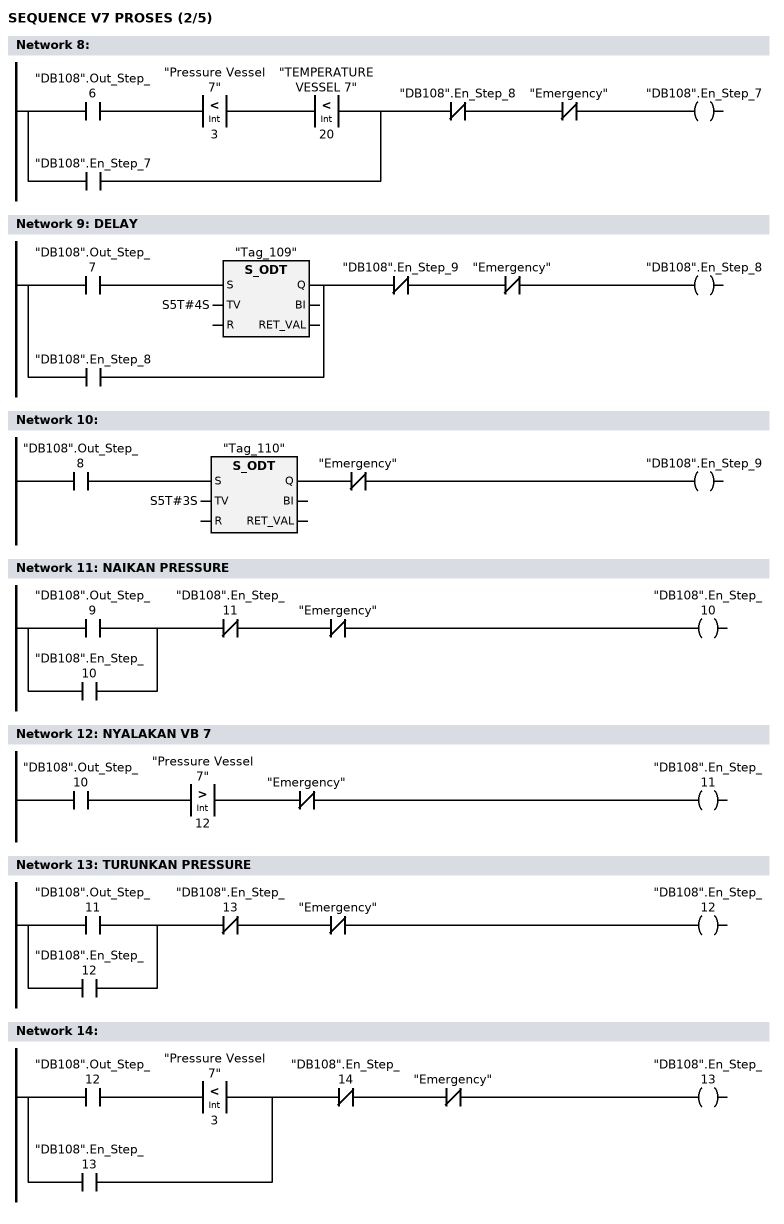
   RUNG wire#powerrail
      Contact( "DB108".Out_Step_6 )
      { S7_Templates := "SrcType := Int" } LT_Contact(in1 := "Pressure Vessel 7", in2 := 3)
      { S7_Templates := "SrcType := Int" } LT_Contact(in1 := "TEMPERATURE VESSEL 7", in2 := 20)
      wire#w1
      I_Contact( "DB108".En_Step_8 )
      I_Contact( "Emergency" )
      Coil( "DB108".En_Step_7 )
   END_RUNG
   RUNG wire#powerrail
      Contact( "DB108".En_Step_7 )
   END_RUNG wire#w1
   // the same network as SCL:
   "DB108".En_Step_7 := (("DB108".Out_Step_6 AND ("Pressure Vessel 7" < 3) AND ("TEMPERATURE VESSEL 7" < 20)) OR "DB108".En_Step_7) AND NOT "DB108".En_Step_8 AND NOT "Emergency";
END_REGION

REGION Network 9: DELAY
   RUNG wire#powerrail
      Contact( "DB108".Out_Step_7 )
      S_ODT(T_NO := "Tag_109", TV := S5T#4S, R :=, BI =>, RET_VAL =>)
      wire#w1
      I_Contact( "DB108".En_Step_9 )
      I_Contact( "Emergency" )
      Coil( "DB108".En_Step_8 )
   END_RUNG
   RUNG wire#powerrail
      Contact( "DB108".En_Step_8 )
   END_RUNG wire#w1
   // the same network as SCL:
   #_s5time1 := S_ODT(T_NO := "Tag_109", S := "DB108".Out_Step_7, TV := S5T#4S, Q => #_w1);
   "DB108".En_Step_8 := (#_w1 OR "DB108".En_Step_8) AND NOT "DB108".En_Step_9 AND NOT "Emergency";
END_REGION

REGION Network 10
   RUNG wire#powerrail
      Contact( "DB108".Out_Step_8 )
      S_ODT(T_NO := "Tag_110", TV := S5T#3S, R :=, BI =>, RET_VAL =>)
      I_Contact( "Emergency" )
      Coil( "DB108".En_Step_9 )
   END_RUNG
   // the same network as SCL:
   #_s5time1 := S_ODT(T_NO := "Tag_110", S := "DB108".Out_Step_8, TV := S5T#3S, Q => #_w1);
   "DB108".En_Step_9 := #_w1 AND NOT "Emergency";
END_REGION

REGION Network 11: NAIKAN PRESSURE
   RUNG wire#powerrail
      Contact( "DB108".Out_Step_9 )
      wire#w1
      I_Contact( "DB108".En_Step_11 )
      I_Contact( "Emergency" )
      Coil( "DB108".En_Step_10 )
   END_RUNG
   RUNG wire#powerrail
      Contact( "DB108".En_Step_10 )
   END_RUNG wire#w1
   // the same network as SCL:
   "DB108".En_Step_10 := ("DB108".Out_Step_9 OR "DB108".En_Step_10) AND NOT "DB108".En_Step_11 AND NOT "Emergency";
END_REGION

REGION Network 12: NYALAKAN VB 7
   RUNG wire#powerrail
      Contact( "DB108".Out_Step_10 )
      { S7_Templates := "SrcType := Int" } GT_Contact(in1 := "Pressure Vessel 7", in2 := 12)
      I_Contact( "Emergency" )
      Coil( "DB108".En_Step_11 )
   END_RUNG
   // the same network as SCL:
   "DB108".En_Step_11 := "DB108".Out_Step_10 AND ("Pressure Vessel 7" > 12) AND NOT "Emergency";
END_REGION

REGION Network 13: TURUNKAN PRESSURE
   RUNG wire#powerrail
      Contact( "DB108".Out_Step_11 )
      wire#w1
      I_Contact( "DB108".En_Step_13 )
      I_Contact( "Emergency" )
      Coil( "DB108".En_Step_12 )
   END_RUNG
   RUNG wire#powerrail
      Contact( "DB108".En_Step_12 )
   END_RUNG wire#w1
   // the same network as SCL:
   "DB108".En_Step_12 := ("DB108".Out_Step_11 OR "DB108".En_Step_12) AND NOT "DB108".En_Step_13 AND NOT "Emergency";
END_REGION

REGION Network 14
   RUNG wire#powerrail
      Contact( "DB108".Out_Step_12 )
      { S7_Templates := "SrcType := Int" } LT_Contact(in1 := "Pressure Vessel 7", in2 := 3)
      wire#w1
      I_Contact( "DB108".En_Step_14 )
      I_Contact( "Emergency" )
      Coil( "DB108".En_Step_13 )
   END_RUNG
   RUNG wire#powerrail
      Contact( "DB108".En_Step_13 )
   END_RUNG wire#w1
   // the same network as SCL:
   "DB108".En_Step_13 := (("DB108".Out_Step_12 AND ("Pressure Vessel 7" < 3)) OR "DB108".En_Step_13) AND NOT "DB108".En_Step_14 AND NOT "Emergency";
END_REGION

REGION Network 15
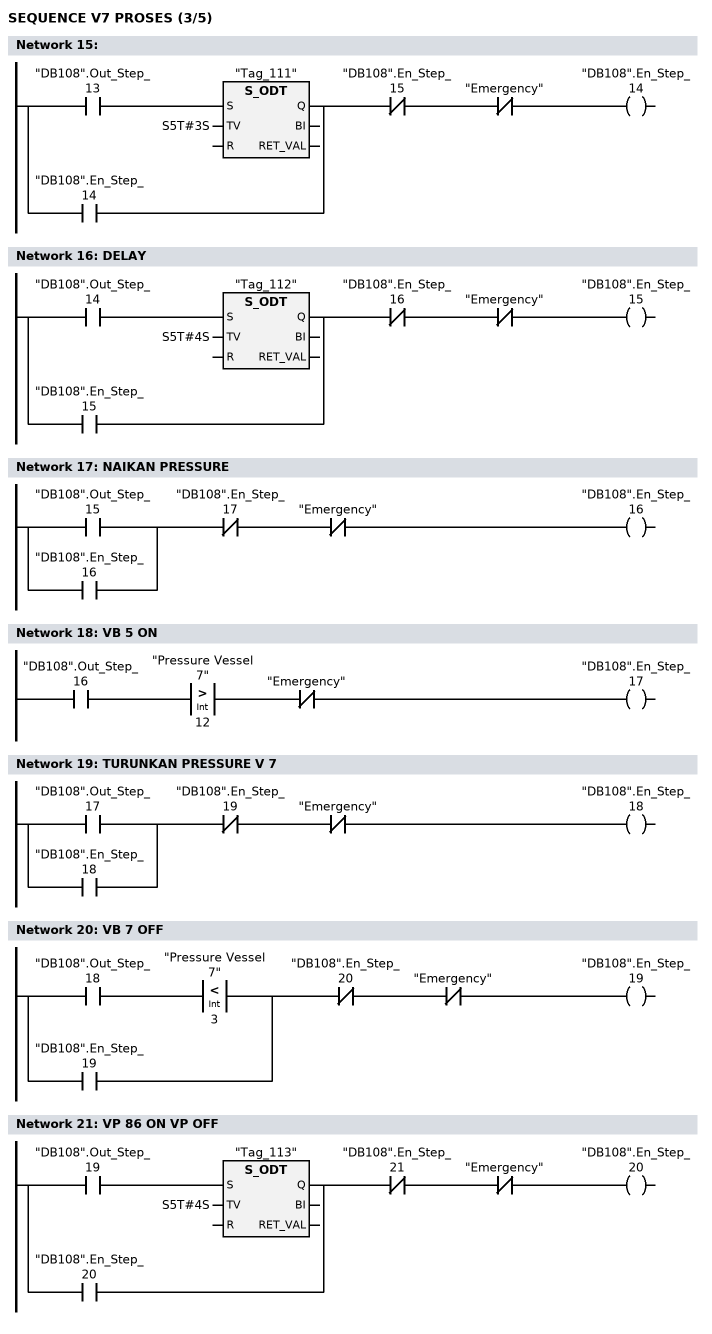
   RUNG wire#powerrail
      Contact( "DB108".Out_Step_13 )
      S_ODT(T_NO := "Tag_111", TV := S5T#3S, R :=, BI =>, RET_VAL =>)
      wire#w1
      I_Contact( "DB108".En_Step_15 )
      I_Contact( "Emergency" )
      Coil( "DB108".En_Step_14 )
   END_RUNG
   RUNG wire#powerrail
      Contact( "DB108".En_Step_14 )
   END_RUNG wire#w1
   // the same network as SCL:
   #_s5time1 := S_ODT(T_NO := "Tag_111", S := "DB108".Out_Step_13, TV := S5T#3S, Q => #_w1);
   "DB108".En_Step_14 := (#_w1 OR "DB108".En_Step_14) AND NOT "DB108".En_Step_15 AND NOT "Emergency";
END_REGION

REGION Network 16: DELAY
   RUNG wire#powerrail
      Contact( "DB108".Out_Step_14 )
      S_ODT(T_NO := "Tag_112", TV := S5T#4S, R :=, BI =>, RET_VAL =>)
      wire#w1
      I_Contact( "DB108".En_Step_16 )
      I_Contact( "Emergency" )
      Coil( "DB108".En_Step_15 )
   END_RUNG
   RUNG wire#powerrail
      Contact( "DB108".En_Step_15 )
   END_RUNG wire#w1
   // the same network as SCL:
   #_s5time1 := S_ODT(T_NO := "Tag_112", S := "DB108".Out_Step_14, TV := S5T#4S, Q => #_w1);
   "DB108".En_Step_15 := (#_w1 OR "DB108".En_Step_15) AND NOT "DB108".En_Step_16 AND NOT "Emergency";
END_REGION

REGION Network 17: NAIKAN PRESSURE
   RUNG wire#powerrail
      Contact( "DB108".Out_Step_15 )
      wire#w1
      I_Contact( "DB108".En_Step_17 )
      I_Contact( "Emergency" )
      Coil( "DB108".En_Step_16 )
   END_RUNG
   RUNG wire#powerrail
      Contact( "DB108".En_Step_16 )
   END_RUNG wire#w1
   // the same network as SCL:
   "DB108".En_Step_16 := ("DB108".Out_Step_15 OR "DB108".En_Step_16) AND NOT "DB108".En_Step_17 AND NOT "Emergency";
END_REGION

REGION Network 18: VB 5 ON
   RUNG wire#powerrail
      Contact( "DB108".Out_Step_16 )
      { S7_Templates := "SrcType := Int" } GT_Contact(in1 := "Pressure Vessel 7", in2 := 12)
      I_Contact( "Emergency" )
      Coil( "DB108".En_Step_17 )
   END_RUNG
   // the same network as SCL:
   "DB108".En_Step_17 := "DB108".Out_Step_16 AND ("Pressure Vessel 7" > 12) AND NOT "Emergency";
END_REGION

REGION Network 19: TURUNKAN PRESSURE V 7
   RUNG wire#powerrail
      Contact( "DB108".Out_Step_17 )
      wire#w1
      I_Contact( "DB108".En_Step_19 )
      I_Contact( "Emergency" )
      Coil( "DB108".En_Step_18 )
   END_RUNG
   RUNG wire#powerrail
      Contact( "DB108".En_Step_18 )
   END_RUNG wire#w1
   // the same network as SCL:
   "DB108".En_Step_18 := ("DB108".Out_Step_17 OR "DB108".En_Step_18) AND NOT "DB108".En_Step_19 AND NOT "Emergency";
END_REGION

REGION Network 20: VB 7 OFF
   RUNG wire#powerrail
      Contact( "DB108".Out_Step_18 )
      { S7_Templates := "SrcType := Int" } LT_Contact(in1 := "Pressure Vessel 7", in2 := 3)
      wire#w1
      I_Contact( "DB108".En_Step_20 )
      I_Contact( "Emergency" )
      Coil( "DB108".En_Step_19 )
   END_RUNG
   RUNG wire#powerrail
      Contact( "DB108".En_Step_19 )
   END_RUNG wire#w1
   // the same network as SCL:
   "DB108".En_Step_19 := (("DB108".Out_Step_18 AND ("Pressure Vessel 7" < 3)) OR "DB108".En_Step_19) AND NOT "DB108".En_Step_20 AND NOT "Emergency";
END_REGION

REGION Network 21: VP 86 ON VP OFF
   RUNG wire#powerrail
      Contact( "DB108".Out_Step_19 )
      S_ODT(T_NO := "Tag_113", TV := S5T#4S, R :=, BI =>, RET_VAL =>)
      wire#w1
      I_Contact( "DB108".En_Step_21 )
      I_Contact( "Emergency" )
      Coil( "DB108".En_Step_20 )
   END_RUNG
   RUNG wire#powerrail
      Contact( "DB108".En_Step_20 )
   END_RUNG wire#w1
   // the same network as SCL:
   #_s5time1 := S_ODT(T_NO := "Tag_113", S := "DB108".Out_Step_19, TV := S5T#4S, Q => #_w1);
   "DB108".En_Step_20 := (#_w1 OR "DB108".En_Step_20) AND NOT "DB108".En_Step_21 AND NOT "Emergency";
END_REGION

REGION Network 22: VP 86 OFF VP 87 ON
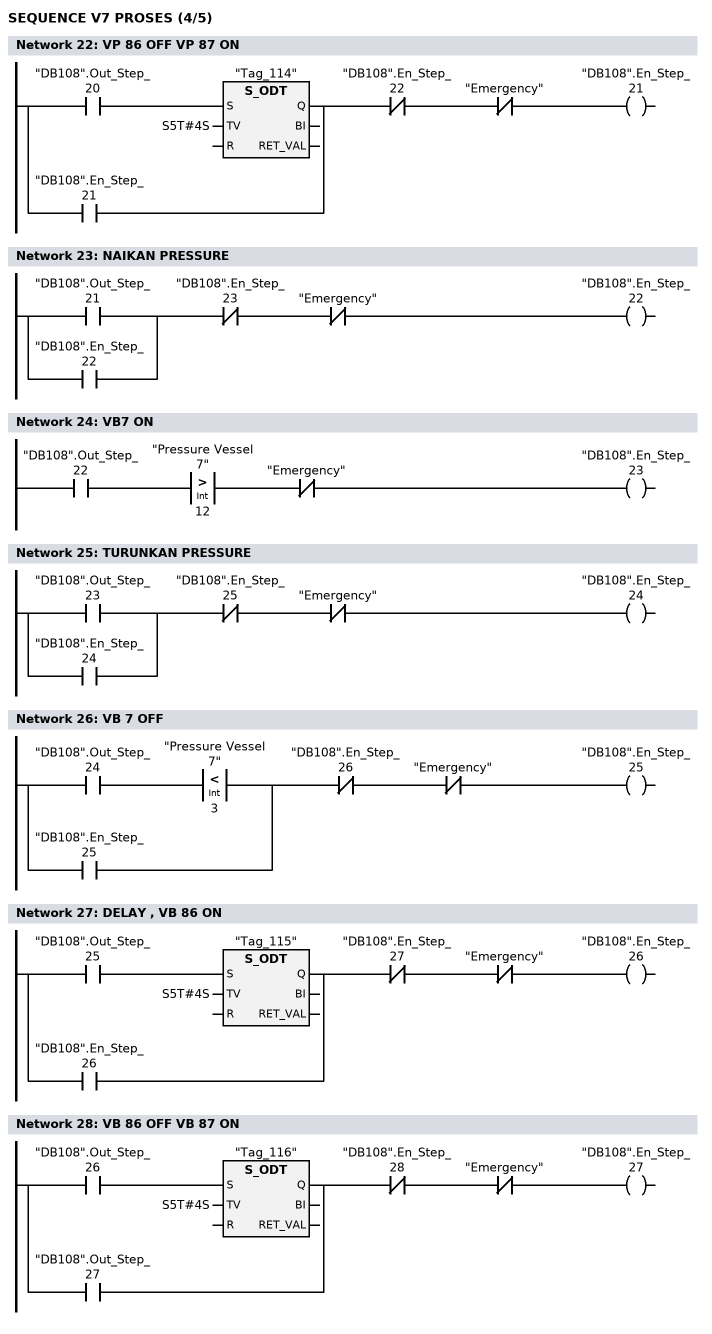
   RUNG wire#powerrail
      Contact( "DB108".Out_Step_20 )
      S_ODT(T_NO := "Tag_114", TV := S5T#4S, R :=, BI =>, RET_VAL =>)
      wire#w1
      I_Contact( "DB108".En_Step_22 )
      I_Contact( "Emergency" )
      Coil( "DB108".En_Step_21 )
   END_RUNG
   RUNG wire#powerrail
      Contact( "DB108".En_Step_21 )
   END_RUNG wire#w1
   // the same network as SCL:
   #_s5time1 := S_ODT(T_NO := "Tag_114", S := "DB108".Out_Step_20, TV := S5T#4S, Q => #_w1);
   "DB108".En_Step_21 := (#_w1 OR "DB108".En_Step_21) AND NOT "DB108".En_Step_22 AND NOT "Emergency";
END_REGION

REGION Network 23: NAIKAN PRESSURE
   RUNG wire#powerrail
      Contact( "DB108".Out_Step_21 )
      wire#w1
      I_Contact( "DB108".En_Step_23 )
      I_Contact( "Emergency" )
      Coil( "DB108".En_Step_22 )
   END_RUNG
   RUNG wire#powerrail
      Contact( "DB108".En_Step_22 )
   END_RUNG wire#w1
   // the same network as SCL:
   "DB108".En_Step_22 := ("DB108".Out_Step_21 OR "DB108".En_Step_22) AND NOT "DB108".En_Step_23 AND NOT "Emergency";
END_REGION

REGION Network 24: VB7 ON
   RUNG wire#powerrail
      Contact( "DB108".Out_Step_22 )
      { S7_Templates := "SrcType := Int" } GT_Contact(in1 := "Pressure Vessel 7", in2 := 12)
      I_Contact( "Emergency" )
      Coil( "DB108".En_Step_23 )
   END_RUNG
   // the same network as SCL:
   "DB108".En_Step_23 := "DB108".Out_Step_22 AND ("Pressure Vessel 7" > 12) AND NOT "Emergency";
END_REGION

REGION Network 25: TURUNKAN PRESSURE
   RUNG wire#powerrail
      Contact( "DB108".Out_Step_23 )
      wire#w1
      I_Contact( "DB108".En_Step_25 )
      I_Contact( "Emergency" )
      Coil( "DB108".En_Step_24 )
   END_RUNG
   RUNG wire#powerrail
      Contact( "DB108".En_Step_24 )
   END_RUNG wire#w1
   // the same network as SCL:
   "DB108".En_Step_24 := ("DB108".Out_Step_23 OR "DB108".En_Step_24) AND NOT "DB108".En_Step_25 AND NOT "Emergency";
END_REGION

REGION Network 26: VB 7 OFF
   RUNG wire#powerrail
      Contact( "DB108".Out_Step_24 )
      { S7_Templates := "SrcType := Int" } LT_Contact(in1 := "Pressure Vessel 7", in2 := 3)
      wire#w1
      I_Contact( "DB108".En_Step_26 )
      I_Contact( "Emergency" )
      Coil( "DB108".En_Step_25 )
   END_RUNG
   RUNG wire#powerrail
      Contact( "DB108".En_Step_25 )
   END_RUNG wire#w1
   // the same network as SCL:
   "DB108".En_Step_25 := (("DB108".Out_Step_24 AND ("Pressure Vessel 7" < 3)) OR "DB108".En_Step_25) AND NOT "DB108".En_Step_26 AND NOT "Emergency";
END_REGION

REGION Network 27: DELAY , VB 86 ON
   RUNG wire#powerrail
      Contact( "DB108".Out_Step_25 )
      S_ODT(T_NO := "Tag_115", TV := S5T#4S, R :=, BI =>, RET_VAL =>)
      wire#w1
      I_Contact( "DB108".En_Step_27 )
      I_Contact( "Emergency" )
      Coil( "DB108".En_Step_26 )
   END_RUNG
   RUNG wire#powerrail
      Contact( "DB108".En_Step_26 )
   END_RUNG wire#w1
   // the same network as SCL:
   #_s5time1 := S_ODT(T_NO := "Tag_115", S := "DB108".Out_Step_25, TV := S5T#4S, Q => #_w1);
   "DB108".En_Step_26 := (#_w1 OR "DB108".En_Step_26) AND NOT "DB108".En_Step_27 AND NOT "Emergency";
END_REGION

REGION Network 28: VB 86 OFF VB 87 ON
   RUNG wire#powerrail
      Contact( "DB108".Out_Step_26 )
      S_ODT(T_NO := "Tag_116", TV := S5T#4S, R :=, BI =>, RET_VAL =>)
      wire#w1
      I_Contact( "DB108".En_Step_28 )
      I_Contact( "Emergency" )
      Coil( "DB108".En_Step_27 )
   END_RUNG
   RUNG wire#powerrail
      Contact( "DB108".Out_Step_27 )
   END_RUNG wire#w1
   // the same network as SCL:
   #_s5time1 := S_ODT(T_NO := "Tag_116", S := "DB108".Out_Step_26, TV := S5T#4S, Q => #_w1);
   "DB108".En_Step_27 := (#_w1 OR "DB108".Out_Step_27) AND NOT "DB108".En_Step_28 AND NOT "Emergency";
END_REGION

REGION Network 29
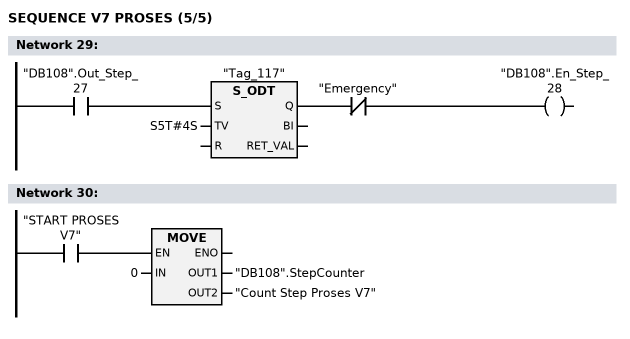
   RUNG wire#powerrail
      Contact( "DB108".Out_Step_27 )
      S_ODT(T_NO := "Tag_117", TV := S5T#4S, R :=, BI =>, RET_VAL =>)
      I_Contact( "Emergency" )
      Coil( "DB108".En_Step_28 )
   END_RUNG
   // the same network as SCL:
   #_s5time1 := S_ODT(T_NO := "Tag_117", S := "DB108".Out_Step_27, TV := S5T#4S, Q => #_w1);
   "DB108".En_Step_28 := #_w1 AND NOT "Emergency";
END_REGION

REGION Network 30
   RUNG wire#powerrail
      Contact( "START PROSES V7" )
      Move(in := 0, out1 => "DB108".StepCounter, out2 => "Count Step Proses V7")
   END_RUNG
   // the same network as SCL:
   IF "START PROSES V7" THEN
       "DB108".StepCounter := 0;
       "Count Step Proses V7" := 0;
   END_IF;
END_REGION
END_FUNCTION

FUNCTION "SEQUENCE V2 PREPARATION" : Void   // FC23, LAD
{ S7_Optimized_Access := 'TRUE' }
VERSION : 0.1
   VAR_TEMP   // added for the SCL form of the ladder/FBD networks
      _w1 : Bool;
      _s5time1 : S5Time;
      _w2 : Bool;
      _s5time2 : S5Time;
   END_VAR
BEGIN

REGION Network 1: Start Preparation
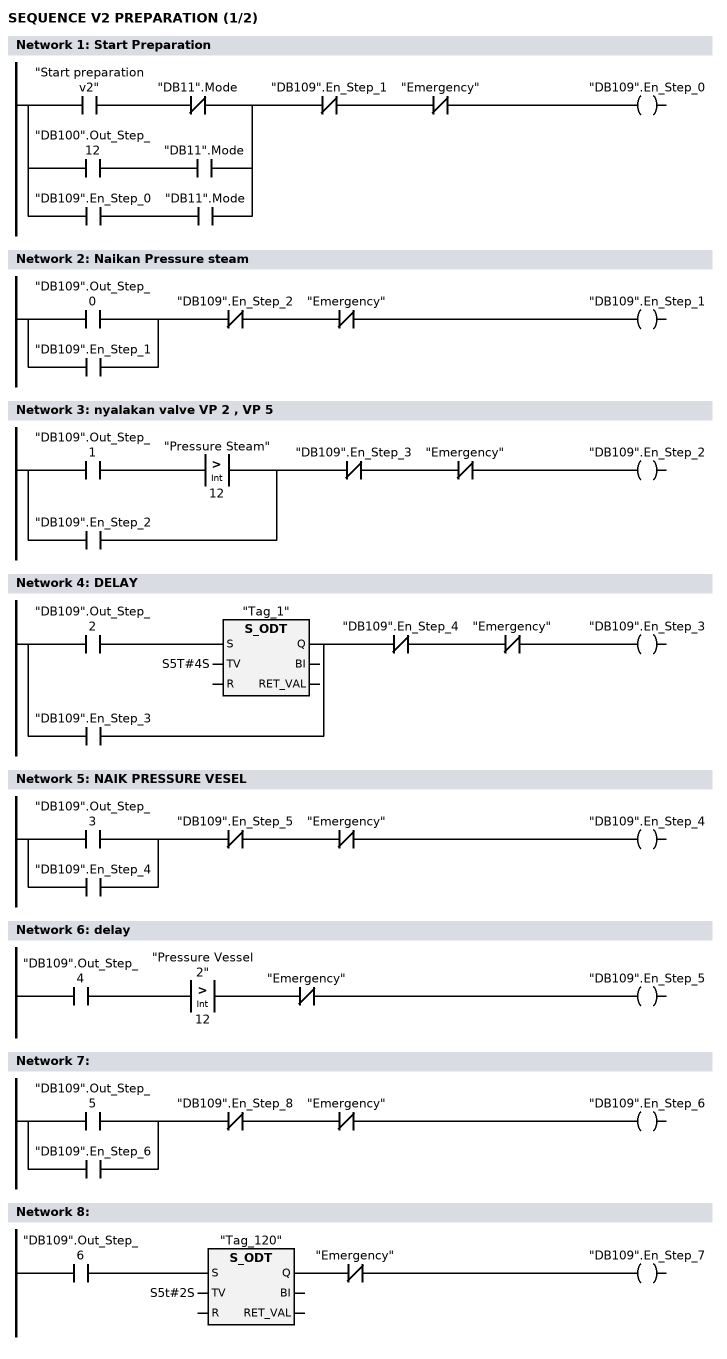
   RUNG wire#powerrail
      Contact( "Start preparation v2" )
      I_Contact( "DB11".Mode )
      wire#w1
      I_Contact( "DB109".En_Step_1 )
      I_Contact( "Emergency" )
      Coil( "DB109".En_Step_0 )
   END_RUNG
   RUNG wire#powerrail
      Contact( "DB100".Out_Step_12 )
      Contact( "DB11".Mode )
   END_RUNG wire#w1
   RUNG wire#powerrail
      Contact( "DB109".En_Step_0 )
      Contact( "DB11".Mode )
   END_RUNG wire#w1
   // the same network as SCL:
   "DB109".En_Step_0 := (("Start preparation v2" AND NOT "DB11".Mode) OR ("DB100".Out_Step_12 AND "DB11".Mode) OR ("DB109".En_Step_0 AND "DB11".Mode)) AND NOT "DB109".En_Step_1 AND NOT "Emergency";
END_REGION

REGION Network 2: Naikan Pressure steam
   RUNG wire#powerrail
      Contact( "DB109".Out_Step_0 )
      wire#w1
      I_Contact( "DB109".En_Step_2 )
      I_Contact( "Emergency" )
      Coil( "DB109".En_Step_1 )
   END_RUNG
   RUNG wire#powerrail
      Contact( "DB109".En_Step_1 )
   END_RUNG wire#w1
   // the same network as SCL:
   "DB109".En_Step_1 := ("DB109".Out_Step_0 OR "DB109".En_Step_1) AND NOT "DB109".En_Step_2 AND NOT "Emergency";
END_REGION

REGION Network 3: nyalakan valve VP 2 , VP 5
   RUNG wire#powerrail
      Contact( "DB109".Out_Step_1 )
      { S7_Templates := "SrcType := Int" } GT_Contact(in1 := "Pressure Steam", in2 := 12)
      wire#w1
      I_Contact( "DB109".En_Step_3 )
      I_Contact( "Emergency" )
      Coil( "DB109".En_Step_2 )
   END_RUNG
   RUNG wire#powerrail
      Contact( "DB109".En_Step_2 )
   END_RUNG wire#w1
   // the same network as SCL:
   "DB109".En_Step_2 := (("DB109".Out_Step_1 AND ("Pressure Steam" > 12)) OR "DB109".En_Step_2) AND NOT "DB109".En_Step_3 AND NOT "Emergency";
END_REGION

REGION Network 4: DELAY
   RUNG wire#powerrail
      Contact( "DB109".Out_Step_2 )
      S_ODT(T_NO := "Tag_1", TV := S5T#4S, R :=, BI =>, RET_VAL =>)
      wire#w1
      I_Contact( "DB109".En_Step_4 )
      I_Contact( "Emergency" )
      Coil( "DB109".En_Step_3 )
   END_RUNG
   RUNG wire#powerrail
      Contact( "DB109".En_Step_3 )
   END_RUNG wire#w1
   // the same network as SCL:
   #_s5time1 := S_ODT(T_NO := "Tag_1", S := "DB109".Out_Step_2, TV := S5T#4S, Q => #_w1);
   "DB109".En_Step_3 := (#_w1 OR "DB109".En_Step_3) AND NOT "DB109".En_Step_4 AND NOT "Emergency";
END_REGION

REGION Network 5: NAIK PRESSURE VESEL
   RUNG wire#powerrail
      Contact( "DB109".Out_Step_3 )
      wire#w1
      I_Contact( "DB109".En_Step_5 )
      I_Contact( "Emergency" )
      Coil( "DB109".En_Step_4 )
   END_RUNG
   RUNG wire#powerrail
      Contact( "DB109".En_Step_4 )
   END_RUNG wire#w1
   // the same network as SCL:
   "DB109".En_Step_4 := ("DB109".Out_Step_3 OR "DB109".En_Step_4) AND NOT "DB109".En_Step_5 AND NOT "Emergency";
END_REGION

REGION Network 6: delay
   RUNG wire#powerrail
      Contact( "DB109".Out_Step_4 )
      { S7_Templates := "SrcType := Int" } GT_Contact(in1 := "Pressure Vessel 2", in2 := 12)
      I_Contact( "Emergency" )
      Coil( "DB109".En_Step_5 )
   END_RUNG
   // the same network as SCL:
   "DB109".En_Step_5 := "DB109".Out_Step_4 AND ("Pressure Vessel 2" > 12) AND NOT "Emergency";
END_REGION

REGION Network 7
   RUNG wire#powerrail
      Contact( "DB109".Out_Step_5 )
      wire#w1
      I_Contact( "DB109".En_Step_8 )
      I_Contact( "Emergency" )
      Coil( "DB109".En_Step_6 )
   END_RUNG
   RUNG wire#powerrail
      Contact( "DB109".En_Step_6 )
   END_RUNG wire#w1
   // the same network as SCL:
   "DB109".En_Step_6 := ("DB109".Out_Step_5 OR "DB109".En_Step_6) AND NOT "DB109".En_Step_8 AND NOT "Emergency";
END_REGION

REGION Network 8
   RUNG wire#powerrail
      Contact( "DB109".Out_Step_6 )
      S_ODT(T_NO := "Tag_120", TV := S5t#2S, R :=, BI =>, RET_VAL =>)
      I_Contact( "Emergency" )
      Coil( "DB109".En_Step_7 )
   END_RUNG
   // the same network as SCL:
   #_s5time1 := S_ODT(T_NO := "Tag_120", S := "DB109".Out_Step_6, TV := S5t#2S, Q => #_w1);
   "DB109".En_Step_7 := #_w1 AND NOT "Emergency";
END_REGION

REGION Network 9: TURUNKAN PRESSURE
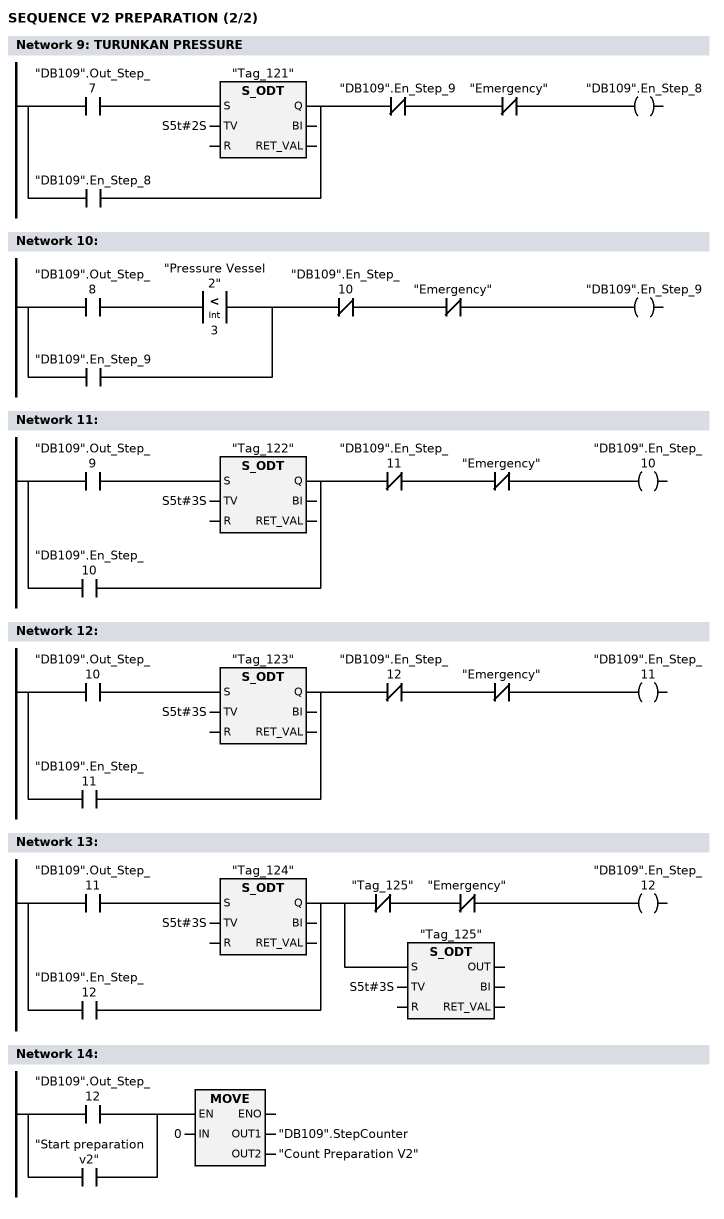
   RUNG wire#powerrail
      Contact( "DB109".Out_Step_7 )
      S_ODT(T_NO := "Tag_121", TV := S5t#2S, R :=, BI =>, RET_VAL =>)
      wire#w1
      I_Contact( "DB109".En_Step_9 )
      I_Contact( "Emergency" )
      Coil( "DB109".En_Step_8 )
   END_RUNG
   RUNG wire#powerrail
      Contact( "DB109".En_Step_8 )
   END_RUNG wire#w1
   // the same network as SCL:
   #_s5time1 := S_ODT(T_NO := "Tag_121", S := "DB109".Out_Step_7, TV := S5t#2S, Q => #_w1);
   "DB109".En_Step_8 := (#_w1 OR "DB109".En_Step_8) AND NOT "DB109".En_Step_9 AND NOT "Emergency";
END_REGION

REGION Network 10
   RUNG wire#powerrail
      Contact( "DB109".Out_Step_8 )
      { S7_Templates := "SrcType := Int" } LT_Contact(in1 := "Pressure Vessel 2", in2 := 3)
      wire#w1
      I_Contact( "DB109".En_Step_10 )
      I_Contact( "Emergency" )
      Coil( "DB109".En_Step_9 )
   END_RUNG
   RUNG wire#powerrail
      Contact( "DB109".En_Step_9 )
   END_RUNG wire#w1
   // the same network as SCL:
   "DB109".En_Step_9 := (("DB109".Out_Step_8 AND ("Pressure Vessel 2" < 3)) OR "DB109".En_Step_9) AND NOT "DB109".En_Step_10 AND NOT "Emergency";
END_REGION

REGION Network 11
   RUNG wire#powerrail
      Contact( "DB109".Out_Step_9 )
      S_ODT(T_NO := "Tag_122", TV := S5t#3S, R :=, BI =>, RET_VAL =>)
      wire#w1
      I_Contact( "DB109".En_Step_11 )
      I_Contact( "Emergency" )
      Coil( "DB109".En_Step_10 )
   END_RUNG
   RUNG wire#powerrail
      Contact( "DB109".En_Step_10 )
   END_RUNG wire#w1
   // the same network as SCL:
   #_s5time1 := S_ODT(T_NO := "Tag_122", S := "DB109".Out_Step_9, TV := S5t#3S, Q => #_w1);
   "DB109".En_Step_10 := (#_w1 OR "DB109".En_Step_10) AND NOT "DB109".En_Step_11 AND NOT "Emergency";
END_REGION

REGION Network 12
   RUNG wire#powerrail
      Contact( "DB109".Out_Step_10 )
      S_ODT(T_NO := "Tag_123", TV := S5t#3S, R :=, BI =>, RET_VAL =>)
      wire#w1
      I_Contact( "DB109".En_Step_12 )
      I_Contact( "Emergency" )
      Coil( "DB109".En_Step_11 )
   END_RUNG
   RUNG wire#powerrail
      Contact( "DB109".En_Step_11 )
   END_RUNG wire#w1
   // the same network as SCL:
   #_s5time1 := S_ODT(T_NO := "Tag_123", S := "DB109".Out_Step_10, TV := S5t#3S, Q => #_w1);
   "DB109".En_Step_11 := (#_w1 OR "DB109".En_Step_11) AND NOT "DB109".En_Step_12 AND NOT "Emergency";
END_REGION

REGION Network 13
   RUNG wire#powerrail
      Contact( "DB109".Out_Step_11 )
      S_ODT(T_NO := "Tag_124", TV := S5t#3S, R :=, BI =>, RET_VAL =>)
      wire#w1
      I_Contact( "Tag_125" )
      I_Contact( "Emergency" )
      Coil( "DB109".En_Step_12 )
   END_RUNG
   RUNG wire#powerrail
      Contact( "DB109".En_Step_12 )
   END_RUNG wire#w1
   RUNG wire#w1
      S_ODT(T_NO := "Tag_125", TV := S5t#3S, R :=, BI =>, RET_VAL =>)
   END_RUNG
   // the same network as SCL:
   #_s5time1 := S_ODT(T_NO := "Tag_124", S := "DB109".Out_Step_11, TV := S5t#3S, Q => #_w1);
   #_w2 := #_w1 OR "DB109".En_Step_12;
   "DB109".En_Step_12 := #_w2 AND NOT "Tag_125" AND NOT "Emergency";
   #_s5time2 := S_ODT(T_NO := "Tag_125", S := #_w2, TV := S5t#3S);
END_REGION

REGION Network 14
   RUNG wire#powerrail
      Contact( "DB109".Out_Step_12 )
      wire#w1
      Move(in := 0, out1 => "DB109".StepCounter, out2 => "Count Preparation V2")
   END_RUNG
   RUNG wire#powerrail
      Contact( "Start preparation v2" )
   END_RUNG wire#w1
   // the same network as SCL:
   IF "DB109".Out_Step_12 OR "Start preparation v2" THEN
       "DB109".StepCounter := 0;
       "Count Preparation V2" := 0;
   END_IF;
END_REGION
END_FUNCTION

FUNCTION "VESSEL 2 PREPARATION" : Void   // FC24, LAD
{ S7_Optimized_Access := 'TRUE' }
VERSION : 0.1
   VAR_TEMP   // added for the SCL form of the ladder/FBD networks
      _w1 : Bool;
      _w2 : Bool;
      _w3 : Bool;
      _w4 : Bool;
   END_VAR
BEGIN

REGION Network 1: NAIKAN PRESSURE STEAM
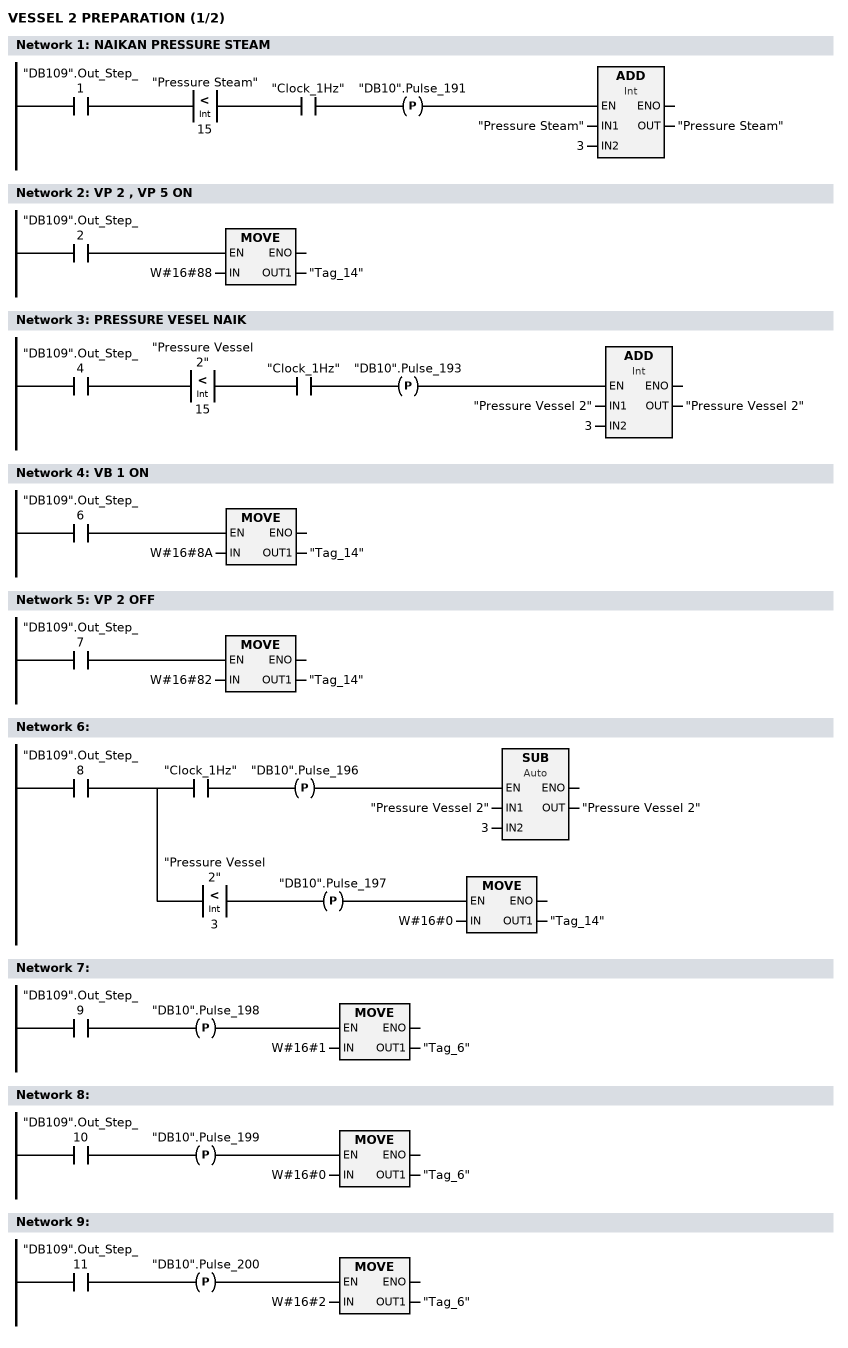
   RUNG wire#powerrail
      Contact( "DB109".Out_Step_1 )
      { S7_Templates := "SrcType := Int" } LT_Contact(in1 := "Pressure Steam", in2 := 15)
      Contact( "Clock_1Hz" )
      P_Trig( "DB10".Pulse_191 )
      { S7_Templates := "SrcType := Int" } Add(in1 := "Pressure Steam", in2 := 3, out => "Pressure Steam")
   END_RUNG
   // the same network as SCL:
   #_w1 := "DB109".Out_Step_1 AND ("Pressure Steam" < 15) AND "Clock_1Hz";
   #_w2 := #_w1 AND NOT "DB10".Pulse_191;   // rising edge
   "DB10".Pulse_191 := #_w1;
   IF #_w2 THEN "Pressure Steam" := "Pressure Steam" + 3; END_IF;
END_REGION

REGION Network 2: VP 2 , VP 5 ON
   RUNG wire#powerrail
      Contact( "DB109".Out_Step_2 )
      Move(in := W#16#88, out1 => "Tag_14")
   END_RUNG
   // the same network as SCL:
   IF "DB109".Out_Step_2 THEN "Tag_14" := W#16#88; END_IF;
END_REGION

REGION Network 3: PRESSURE VESEL NAIK
   RUNG wire#powerrail
      Contact( "DB109".Out_Step_4 )
      { S7_Templates := "SrcType := Int" } LT_Contact(in1 := "Pressure Vessel 2", in2 := 15)
      Contact( "Clock_1Hz" )
      P_Trig( "DB10".Pulse_193 )
      { S7_Templates := "SrcType := Int" } Add(in1 := "Pressure Vessel 2", in2 := 3, out => "Pressure Vessel 2")
   END_RUNG
   // the same network as SCL:
   #_w1 := "DB109".Out_Step_4 AND ("Pressure Vessel 2" < 15) AND "Clock_1Hz";
   #_w2 := #_w1 AND NOT "DB10".Pulse_193;   // rising edge
   "DB10".Pulse_193 := #_w1;
   IF #_w2 THEN "Pressure Vessel 2" := "Pressure Vessel 2" + 3; END_IF;
END_REGION

REGION Network 4: VB 1 ON
   RUNG wire#powerrail
      Contact( "DB109".Out_Step_6 )
      Move(in := W#16#8A, out1 => "Tag_14")
   END_RUNG
   // the same network as SCL:
   IF "DB109".Out_Step_6 THEN "Tag_14" := W#16#8A; END_IF;
END_REGION

REGION Network 5: VP 2 OFF
   RUNG wire#powerrail
      Contact( "DB109".Out_Step_7 )
      Move(in := W#16#82, out1 => "Tag_14")
   END_RUNG
   // the same network as SCL:
   IF "DB109".Out_Step_7 THEN "Tag_14" := W#16#82; END_IF;
END_REGION

REGION Network 6
   RUNG wire#powerrail
      Contact( "DB109".Out_Step_8 )
      wire#w1
      Contact( "Clock_1Hz" )
      P_Trig( "DB10".Pulse_196 )
      Sub(in1 := "Pressure Vessel 2", in2 := 3, out => "Pressure Vessel 2")
   END_RUNG
   RUNG wire#w1
      { S7_Templates := "SrcType := Int" } LT_Contact(in1 := "Pressure Vessel 2", in2 := 3)
      P_Trig( "DB10".Pulse_197 )
      Move(in := W#16#0, out1 => "Tag_14")
   END_RUNG
   // the same network as SCL:
   #_w1 := "DB109".Out_Step_8 AND "Clock_1Hz";
   #_w2 := #_w1 AND NOT "DB10".Pulse_196;   // rising edge
   "DB10".Pulse_196 := #_w1;
   IF #_w2 THEN "Pressure Vessel 2" := "Pressure Vessel 2" - 3; END_IF;
   #_w3 := "DB109".Out_Step_8 AND ("Pressure Vessel 2" < 3);
   #_w4 := #_w3 AND NOT "DB10".Pulse_197;   // rising edge
   "DB10".Pulse_197 := #_w3;
   IF #_w4 THEN "Tag_14" := W#16#0; END_IF;
END_REGION

REGION Network 7
   RUNG wire#powerrail
      Contact( "DB109".Out_Step_9 )
      P_Trig( "DB10".Pulse_198 )
      Move(in := W#16#1, out1 => "Tag_6")
   END_RUNG
   // the same network as SCL:
   #_w1 := "DB109".Out_Step_9 AND NOT "DB10".Pulse_198;   // rising edge
   "DB10".Pulse_198 := "DB109".Out_Step_9;
   IF #_w1 THEN "Tag_6" := W#16#1; END_IF;
END_REGION

REGION Network 8
   RUNG wire#powerrail
      Contact( "DB109".Out_Step_10 )
      P_Trig( "DB10".Pulse_199 )
      Move(in := W#16#0, out1 => "Tag_6")
   END_RUNG
   // the same network as SCL:
   #_w1 := "DB109".Out_Step_10 AND NOT "DB10".Pulse_199;   // rising edge
   "DB10".Pulse_199 := "DB109".Out_Step_10;
   IF #_w1 THEN "Tag_6" := W#16#0; END_IF;
END_REGION

REGION Network 9
   RUNG wire#powerrail
      Contact( "DB109".Out_Step_11 )
      P_Trig( "DB10".Pulse_200 )
      Move(in := W#16#2, out1 => "Tag_6")
   END_RUNG
   // the same network as SCL:
   #_w1 := "DB109".Out_Step_11 AND NOT "DB10".Pulse_200;   // rising edge
   "DB10".Pulse_200 := "DB109".Out_Step_11;
   IF #_w1 THEN "Tag_6" := W#16#2; END_IF;
END_REGION

REGION Network 10
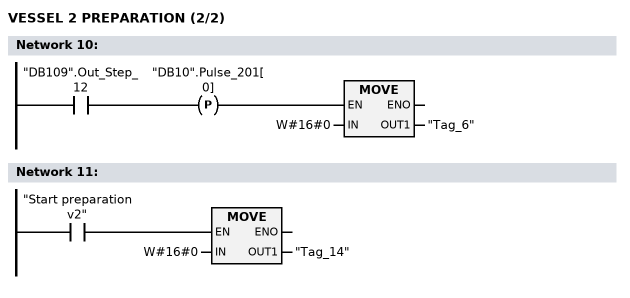
   RUNG wire#powerrail
      Contact( "DB109".Out_Step_12 )
      P_Trig( "DB10".Pulse_201[0] )
      Move(in := W#16#0, out1 => "Tag_6")
   END_RUNG
   // the same network as SCL:
   #_w1 := "DB109".Out_Step_12 AND NOT "DB10".Pulse_201[0];   // rising edge
   "DB10".Pulse_201[0] := "DB109".Out_Step_12;
   IF #_w1 THEN "Tag_6" := W#16#0; END_IF;
END_REGION

REGION Network 11
   RUNG wire#powerrail
      Contact( "Start preparation v2" )
      Move(in := W#16#0, out1 => "Tag_14")
   END_RUNG
   // the same network as SCL:
   IF "Start preparation v2" THEN "Tag_14" := W#16#0; END_IF;
END_REGION
END_FUNCTION

FUNCTION "SEQUENCE V3 PREPARATION" : Void   // FC25, LAD
{ S7_Optimized_Access := 'TRUE' }
VERSION : 0.1
   VAR_TEMP   // added for the SCL form of the ladder/FBD networks
      _w1 : Bool;
      _s5time1 : S5Time;
      _w2 : Bool;
      _s5time2 : S5Time;
   END_VAR
BEGIN

REGION Network 1: Start Preparation